// TIA Portal project "PROJECT_PC_SUT" (V17)

(* hardware
DEVICE "S7-1500/ET200MP station_1"  S7-1500 station
   slot 0: "Rail_0"  Rack  6ES7 590-1***0-0AA0
   slot 1: "PLC_2"  CPU 1513-1 PN  6ES7 513-1AL01-0AB0  V2.9
      slot 3: "CPU display_1"  6ES7591-1AA00-0AA0
      slot 32768: "PROFINET interface_1"  X1
         slot 32769: "Port_1"  X1 P1
         slot 32770: "Port_2"  X1 P2
      slot 34817: "Virtual CP interface port_1"  Virtual CP interface port  Virtual CP interface port
DEVICE "HMI_1"  TP700 Comfort
   slot 0: "HMI_1"  TP700 Comfort  6AV2 124-0GC01-0AX0  17.0.0.0
   slot 1: "HMI_RT_1"  TP700 Comfort  6AV2 124-0GC01-0AX0  17.0.0.0
   slot 5: "HMI_1.IE_CP_1"  PROFINET Interface  17.0.0.0
      slot 1: "PROFINET Interface_1"  PROFINET Interface
         slot 1: "Port_1"  Port
         slot 2: "Port_2"  Port
   slot 7: "HMI_1.MPI/DP_CP_1"  MPI/DP Interface  17.0.0.0
DEVICE "PC-System_1"  SIMATIC PC station
   slot 0: "SIMATIC PC station"  Rail  SIMATIC PC-Station  V1.0
      slot 125: "Stationmanager"  Station_Manager  V6.0.4
   slot 1: "IE general_1"  IE General  IE_CP  V8.2.0
      slot 1: "PROFINET interface"  IEGeneral.Interface.8.2.0
   slot 2: "HMI_RT_2"  WinCC RT Advanced  6AV2 104-0xxxx-xxxx  17.0.0.0
      slot 33792: "Computer interface"  Host interface
*)

// ===== PLC "PLC_2"  CPU 1513-1 PN =====

VAR_GLOBAL   // PLC tag table "Tag_Table"
   "start" AT %I0.1 : Bool;
   "AI1_level_sensor" AT %IW1 : Int;
   "AI2_temp_sensor" AT %IW3 : Int;
   "set_temperature_MW4" AT %MW4 : Int;
   "initial_temperature_MW6" AT %MW6 : Int;
   "set_level_MW2" AT %MW2 : Int;
   "gain" AT %MW8 : Int;
   "valve1" AT %Q0.1 : Bool;
   "valve2" AT %Q0.2 : Bool;
   "valve3" AT %Q0.3 : Bool;
   "valve4" AT %Q0.4 : Bool;
   "valve5" AT %Q0.5 : Bool;
   "mixer_motor" AT %Q0.6 : Bool;
   "AV1" AT %QW2 : Word;
   "AV2" AT %QW4 : Int;
   "compare_level" AT %MD10 : Real;
   "flag1" AT %M22.0 : Bool;
   "compare_bit_for_heating" AT %M22.1 : Bool;
   "set_heating" AT %M22.2 : Bool;
   "flag2" AT %M22.3 : Bool;
   "flag3" AT %M22.4 : Bool;
   "set_cooling" AT %M22.5 : Bool;
   "flag0" AT %M22.6 : Bool;
   "compare_bit_reset" AT %M22.7 : Bool;
   "compare_drain_bit_1" AT %M23.0 : Bool;
   "compare_drain_bit_2" AT %M23.1 : Bool;
   "drain_activation_bit" AT %M23.2 : Bool;
END_VAR

// folder: System blocks/Program resources

DATA_BLOCK "Timer_1"   // DB1
{ S7_Optimized_Access := 'TRUE' }
AUTHOR : Simatic
FAMILY : IEC
NAME : IEC_TMR
VERSION : 1.0
// stored: InstanceOfName IEC_TIMER
"IEC_TIMER"
BEGIN
END_DATA_BLOCK

// folder: (top level)

FUNCTION "compare_level_value" : Void   // FC1, LAD
{ S7_Optimized_Access := 'TRUE' }
VERSION : 0.1
   VAR_INPUT
      set_level_MW2 : Int;
   END_VAR
   VAR_OUTPUT
      compare_level : Real;
   END_VAR
   VAR_TEMP
      hold : Real;
      set_level_convert : Real;
   END_VAR
BEGIN

REGION Network 1: Data type conversion
   // covert set_level_MW2 from INT to REAL
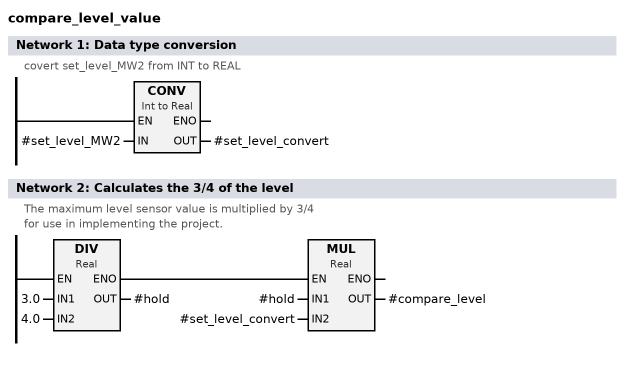
   RUNG wire#powerrail
      { S7_Templates := "[SrcType := Int, DestType := Real]" } Convert(in := #set_level_MW2, out => #set_level_convert)
   END_RUNG
   // the same network as SCL:
   #set_level_convert := INT_TO_REAL(#set_level_MW2);
END_REGION

REGION Network 2: Calculates the 3/4 of the level
   // The maximum level sensor value is multiplied by 3/4
   // for use in implementing the project.
   RUNG wire#powerrail
      { S7_Templates := "SrcType := Real" } Div(in1 := 3.0, in2 := 4.0, out => #hold)
      { S7_Templates := "SrcType := Real" } Mul(in1 := #hold, in2 := #set_level_convert, out => #compare_level)
   END_RUNG
   // the same network as SCL:
   #hold := 3.0 / 4.0;
   #compare_level := #hold * #set_level_convert;
END_REGION
END_FUNCTION

FUNCTION "Filling" : Void   // FC2, LAD
{ S7_Optimized_Access := 'TRUE' }
VERSION : 0.1
   VAR_INPUT
      valve3 : Bool;
      valve4 : Bool;
      valve5 : Bool;
      AI1_level_sensor : Int;
      compare_level : Real;
      set_level_MW2 : Int;
   END_VAR
   VAR_OUTPUT
      valve1 : Bool;
      valve2 : Bool;
      mixer_motor : Bool;
      flag0 : Bool;
   END_VAR
   VAR_TEMP
      level_sensor_conv : Real;
      set_level_converted : Real;
   END_VAR
   VAR_TEMP   // added for the SCL form of the ladder/FBD networks
      _w1 : Bool;
   END_VAR
BEGIN

REGION Network 1: Data type convert
   // A1I_level_sensor data type is converted to Real
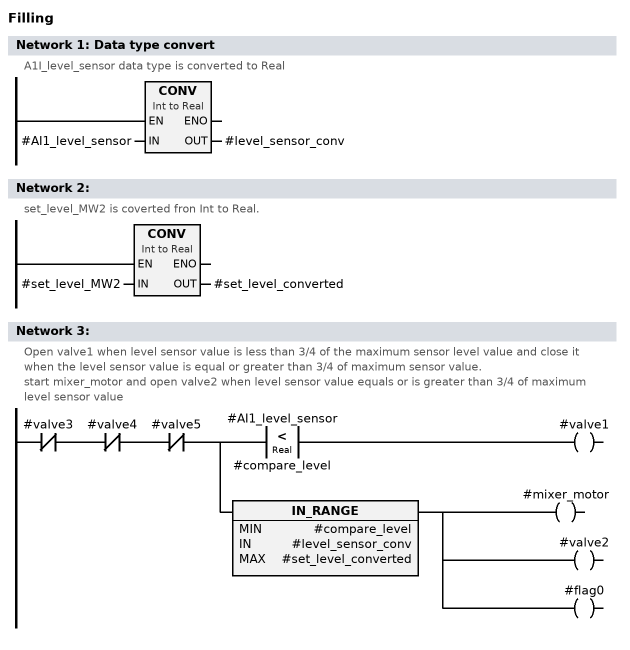
   RUNG wire#powerrail
      { S7_Templates := "[SrcType := Int, DestType := Real]" } Convert(in := #AI1_level_sensor, out => #level_sensor_conv)
   END_RUNG
   // the same network as SCL:
   #level_sensor_conv := INT_TO_REAL(#AI1_level_sensor);
END_REGION

REGION Network 2
   // set_level_MW2 is coverted fron Int to Real.
   RUNG wire#powerrail
      { S7_Templates := "[SrcType := Int, DestType := Real]" } Convert(in := #set_level_MW2, out => #set_level_converted)
   END_RUNG
   // the same network as SCL:
   #set_level_converted := INT_TO_REAL(#set_level_MW2);
END_REGION

REGION Network 3
   // Open valve1 when level sensor value is less than 3/4 of the maximum sensor level value and close it when the level sensor value is equal or greater than 3/4 of maximum sensor value.
   // 
   // start mixer_motor and open valve2 when level sensor value equals or is greater than 3/4 of maximum level sensor value
   RUNG wire#powerrail
      I_Contact( #valve3 )
      I_Contact( #valve4 )
      I_Contact( #valve5 )
      wire#w1
      { S7_Templates := "SrcType := Real" } LT_Contact(in1 := #AI1_level_sensor, in2 := #compare_level)
      Coil( #valve1 )
   END_RUNG
   RUNG wire#w1
      { S7_Templates := "SrcType := Real" } InRange(min := #compare_level, in := #level_sensor_conv, max := #set_level_converted)
      wire#w2
      Coil( #mixer_motor )
   END_RUNG
   RUNG wire#w2
      Coil( #valve2 )
   END_RUNG
   RUNG wire#w2
      Coil( #flag0 )
   END_RUNG
   // the same network as SCL:
   #_w1 := NOT #valve3 AND NOT #valve4 AND NOT #valve5;
   #valve1 := #_w1 AND (#AI1_level_sensor < #compare_level);
   #mixer_motor := #_w1 AND (#compare_level <= #level_sensor_conv) AND (#level_sensor_conv <= #set_level_converted);
   #valve2 := #mixer_motor;
   #flag0 := #mixer_motor;
END_REGION
END_FUNCTION

FUNCTION "P_Controller" : Void   // FC3, LAD
{ S7_Optimized_Access := 'TRUE' }
VERSION : 0.1
// Proportional controller for the system
   VAR_INPUT
      AI2_temp_sensor : Int;
      gain : Int;
      set_temperature_MW4 : Int;
   END_VAR
   VAR_OUTPUT
      AV2 : Int;
   END_VAR
   VAR_TEMP
      error : Int;
      multiply : Real;
      norm_out : Real;
      limit_out : Real;
   END_VAR
BEGIN

REGION Network 1
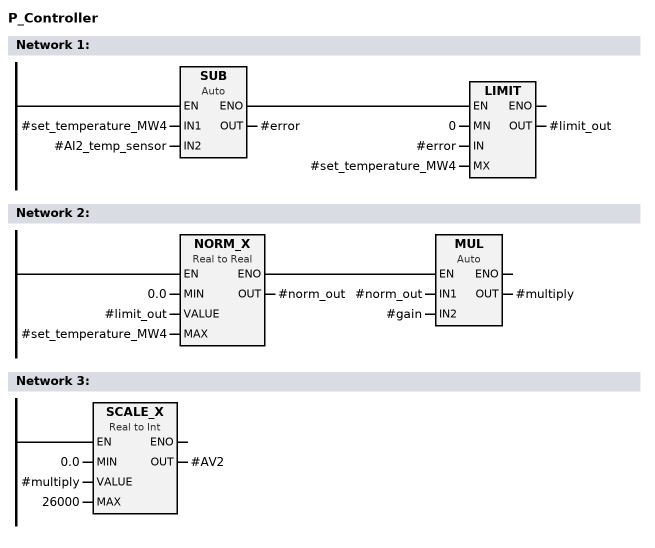
   #error := #set_temperature_MW4 - #AI2_temp_sensor;
   #limit_out := LIMIT(MN := 0, IN := #error, MX := #set_temperature_MW4);
END_REGION

REGION Network 2
   RUNG wire#powerrail
      { S7_Templates := "[SrcType := Real, DestType := Real]" } Normalize(min := 0.0, value := #limit_out, max := #set_temperature_MW4, out => #norm_out)
      Mul(in1 := #norm_out, in2 := #gain, out => #multiply)
   END_RUNG
   // the same network as SCL:
   #norm_out := NORM_X(MIN := 0.0, VALUE := #limit_out, MAX := #set_temperature_MW4);
   #multiply := #norm_out * #gain;
END_REGION

REGION Network 3
   RUNG wire#powerrail
      { S7_Templates := "[SrcType := Real, DestType := Int]" } Scale(min := 0.0, value := #multiply, max := 26000, out => #AV2)
   END_RUNG
   // the same network as SCL:
   #AV2 := SCALE_X(MIN := 0.0, VALUE := #multiply, MAX := 26000);
END_REGION
END_FUNCTION

FUNCTION "heating" : Void   // FC4, LAD
{ S7_Optimized_Access := 'TRUE' }
VERSION : 0.1
   VAR_INPUT
      AI2_temp_sensor : Int;
      valve3 : Bool;
      valve4 : Bool;
      set_temperture_MW4 : Int;
      gain : Int;
   END_VAR
   VAR_OUTPUT
      valve5 : Bool;
      AV2 : Int;
   END_VAR
   VAR_IN_OUT
      trigger_move : Bool;
      flag1 : Bool;
   END_VAR
   VAR_TEMP
      bit_operate : Bool;
   END_VAR
BEGIN

REGION Network 1
   // Reset flag1, which stops mixer_motor and closes valve2 when level sensor value is greater than the set_level sensor value.
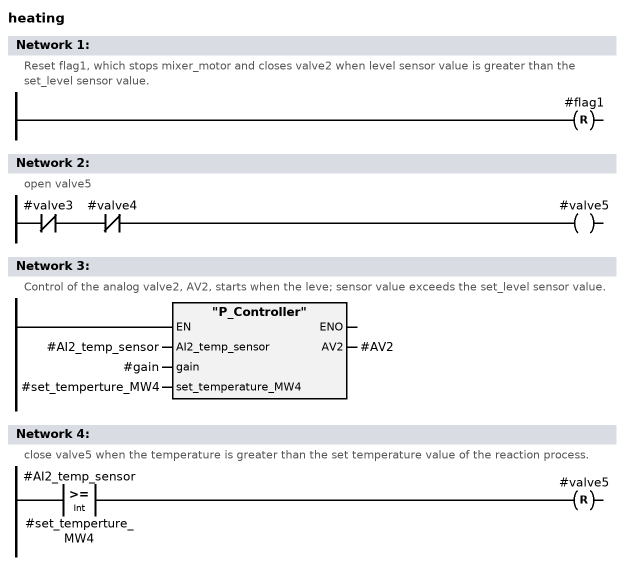
   RUNG wire#powerrail
      R_Coil( #flag1 )
   END_RUNG
   // the same network as SCL:
   #flag1 := FALSE;
END_REGION

REGION Network 2
   // open valve5
   RUNG wire#powerrail
      I_Contact( #valve3 )
      I_Contact( #valve4 )
      Coil( #valve5 )
   END_RUNG
   // the same network as SCL:
   #valve5 := NOT #valve3 AND NOT #valve4;
END_REGION

REGION Network 3
   // Control of the analog valve2, AV2, starts when the leve; sensor value exceeds the set_level sensor value.
   RUNG wire#powerrail
      "P_Controller"(AI2_temp_sensor := #AI2_temp_sensor, gain := #gain, set_temperature_MW4 := #set_temperture_MW4, AV2 => #AV2)
   END_RUNG
   // the same network as SCL:
   "P_Controller"(AI2_temp_sensor := #AI2_temp_sensor,
                  gain := #gain,
                  set_temperature_MW4 := #set_temperture_MW4,
                  AV2 => #AV2);
END_REGION

REGION Network 4
   // close valve5 when the temperature is greater than the set temperature value of the reaction process.
   RUNG wire#powerrail
      { S7_Templates := "SrcType := Int" } GE_Contact(in1 := #AI2_temp_sensor, in2 := #set_temperture_MW4)
      R_Coil( #valve5 )
   END_RUNG
   // the same network as SCL:
   IF #AI2_temp_sensor >= #set_temperture_MW4 THEN #valve5 := FALSE; END_IF;
END_REGION
END_FUNCTION

ORGANIZATION_BLOCK "Main"   // OB1, LAD, ProgramCycle
TITLE = "Main Program Sweep (Cycle)"
{ S7_Optimized_Access := 'TRUE' }
VERSION : 0.1
   VAR_INPUT
      Initial_Call : Bool;   // Initial call of this OB
      Remanence : Bool;   // =True, if remanent data are available
   END_VAR
   VAR_TEMP   // added for the SCL form of the ladder/FBD networks
      _w1 : Bool;
      _w2 : Bool;
      _w3 : Bool;
   END_VAR
BEGIN

REGION Network 1: INITIAL STATE OF THE REACTOR
   // In this block, the compare function is called. This compare function is used to control the mixer and filling processes by comparing the level at which the mixer will be turned on and off, and also when the filling valves will be turned on and off.
   // 
   // Also, we set flag1 in this Network, Flag1 will be used to start the filling phase of the process.
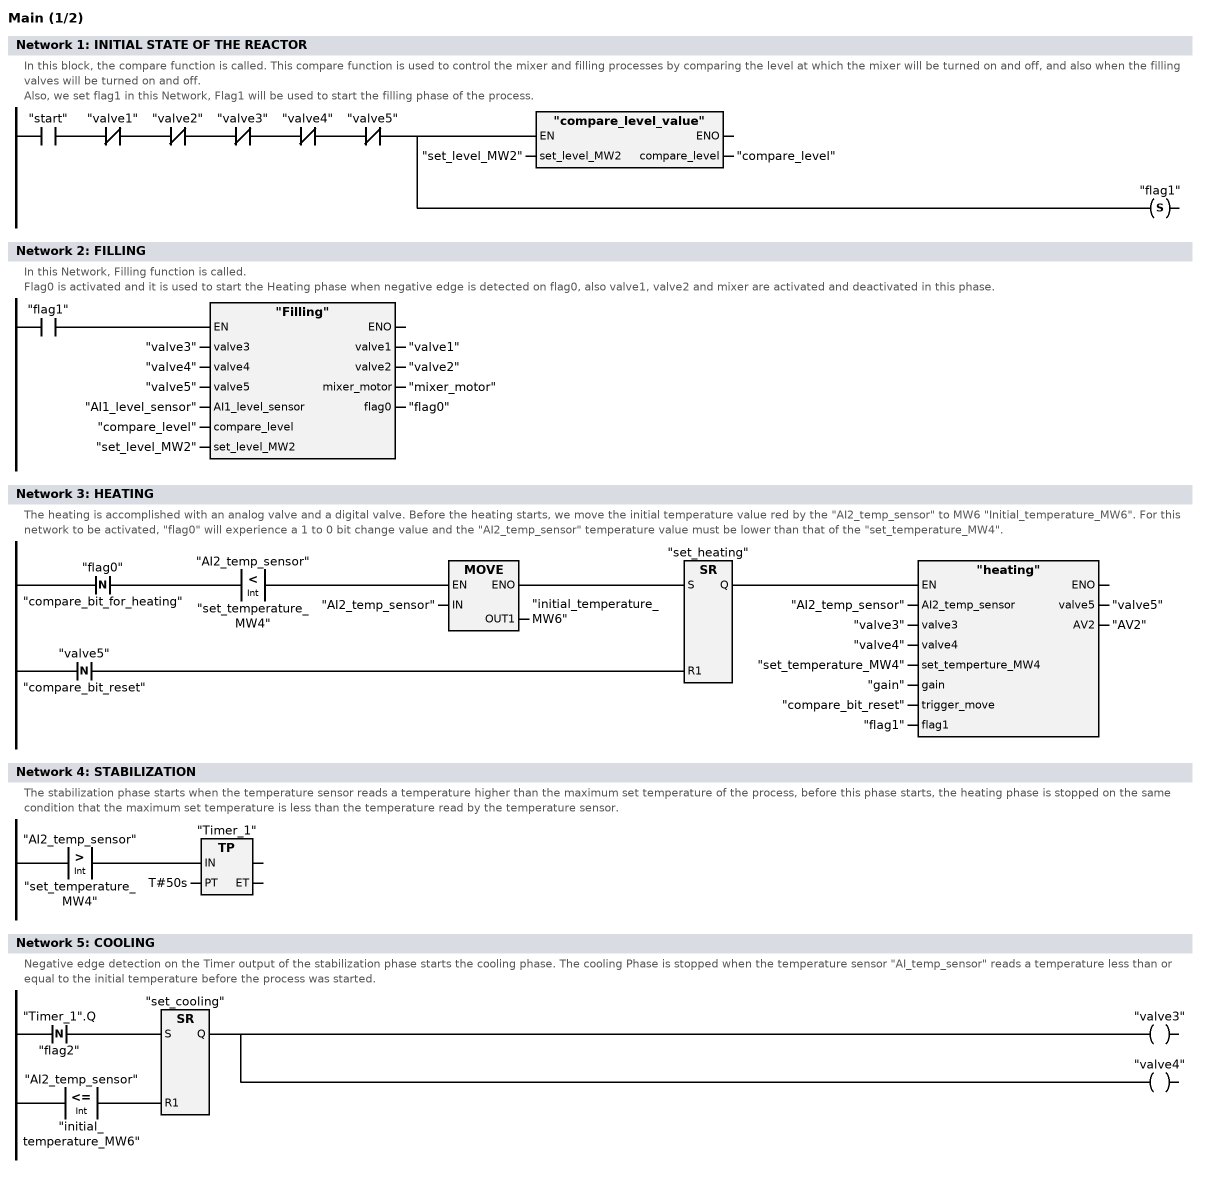
   RUNG wire#powerrail
      Contact( "start" )
      I_Contact( "valve1" )
      I_Contact( "valve2" )
      I_Contact( "valve3" )
      I_Contact( "valve4" )
      I_Contact( "valve5" )
      wire#w1
      "compare_level_value"(set_level_MW2 := "set_level_MW2", compare_level => "compare_level")
   END_RUNG
   RUNG wire#w1
      S_Coil( "flag1" )
   END_RUNG
   // the same network as SCL:
   #_w1 := "start" AND NOT "valve1" AND NOT "valve2" AND NOT "valve3" AND NOT "valve4" AND NOT "valve5";
   IF #_w1 THEN
       "compare_level_value"(set_level_MW2 := "set_level_MW2", compare_level => "compare_level");
       "flag1" := TRUE;
   END_IF;
END_REGION

REGION Network 2: FILLING
   // In this Network, Filling function is called.
   // Flag0 is activated and it is used to start the Heating phase when negative edge is detected on flag0, also valve1, valve2 and mixer are activated and deactivated in this phase.
   RUNG wire#powerrail
      Contact( "flag1" )
      "Filling"(valve3 := "valve3", valve4 := "valve4", valve5 := "valve5", AI1_level_sensor := "AI1_level_sensor", compare_level := "compare_level", set_level_MW2 := "set_level_MW2", valve1 => "valve1", valve2 => "valve2", mixer_motor => "mixer_motor", flag0 => "flag0")
   END_RUNG
   // the same network as SCL:
   IF "flag1" THEN
       "Filling"(valve3 := "valve3",
                 valve4 := "valve4",
                 valve5 := "valve5",
                 AI1_level_sensor := "AI1_level_sensor",
                 compare_level := "compare_level",
                 set_level_MW2 := "set_level_MW2",
                 valve1 => "valve1",
                 valve2 => "valve2",
                 mixer_motor => "mixer_motor",
                 flag0 => "flag0");
   END_IF;
END_REGION

REGION Network 3: HEATING
   // The heating is accomplished with an analog valve and a digital valve. Before the heating starts, we move the initial temperature value red by the "AI2_temp_sensor" to MW6 "Initial_temperature_MW6". For this network to be activated, "flag0" will experience a 1 to 0 bit change value and the "AI2_temp_sensor" temperature value must be lower than that of the "set_temperature_MW4".
   RUNG wire#powerrail
      N_Contact(operand := "flag0", bit := "compare_bit_for_heating")
      { S7_Templates := "SrcType := Int" } LT_Contact(in1 := "AI2_temp_sensor", in2 := "set_temperature_MW4")
      Move(in := "AI2_temp_sensor", out1 => "initial_temperature_MW6")
      S_SR(operand := "set_heating", r1 := wire#w1)
      "heating"(AI2_temp_sensor := "AI2_temp_sensor", valve3 := "valve3", valve4 := "valve4", set_temperture_MW4 := "set_temperature_MW4", gain := "gain", trigger_move := "compare_bit_reset", flag1 := "flag1", valve5 => "valve5", AV2 => "AV2")
   END_RUNG
   RUNG wire#powerrail
      N_Contact(operand := "valve5", bit := "compare_bit_reset")
   END_RUNG wire#w1
   // the same network as SCL:
   #_w1 := NOT "flag0" AND "compare_bit_for_heating";   // falling edge of "flag0"
   "compare_bit_for_heating" := "flag0";
   #_w2 := #_w1 AND ("AI2_temp_sensor" < "set_temperature_MW4");
   IF #_w2 THEN "initial_temperature_MW6" := "AI2_temp_sensor"; END_IF;
   #_w3 := NOT "valve5" AND "compare_bit_reset";   // falling edge of "valve5"
   "compare_bit_reset" := "valve5";
   IF #_w2 THEN
       "set_heating" := TRUE;   // SR flip-flop
   END_IF;
   IF #_w3 THEN "set_heating" := FALSE; END_IF;
   IF "set_heating" THEN
       "heating"(AI2_temp_sensor := "AI2_temp_sensor",
                 valve3 := "valve3",
                 valve4 := "valve4",
                 set_temperture_MW4 := "set_temperature_MW4",
                 gain := "gain",
                 trigger_move := "compare_bit_reset",
                 flag1 := "flag1",
                 valve5 => "valve5",
                 AV2 => "AV2");
   END_IF;
END_REGION

REGION Network 4: STABILIZATION
   // The stabilization phase starts when the temperature sensor reads a temperature higher than the maximum set temperature of the process, before this phase starts, the heating phase is stopped on the same condition that the maximum set temperature is less than the temperature read by the temperature sensor.
   "Timer_1".TP(IN := "AI2_temp_sensor" > "set_temperature_MW4", PT := T#50s);
END_REGION

REGION Network 5: COOLING
   // Negative edge detection on the Timer output of the stabilization phase starts the cooling phase. The cooling Phase is stopped when the temperature sensor "AI_temp_sensor" reads a temperature less than or equal to the initial temperature before the process was started.
   RUNG wire#powerrail
      N_Contact(operand := "Timer_1".Q, bit := "flag2")
      S_SR(operand := "set_cooling", r1 := wire#w1)
      wire#w2
      Coil( "valve3" )
   END_RUNG
   RUNG wire#powerrail
      { S7_Templates := "SrcType := Int" } LE_Contact(in1 := "AI2_temp_sensor", in2 := "initial_temperature_MW6")
   END_RUNG wire#w1
   RUNG wire#w2
      Coil( "valve4" )
   END_RUNG
   // the same network as SCL:
   #_w1 := NOT "Timer_1".Q AND "flag2";   // falling edge of "Timer_1".Q
   "flag2" := "Timer_1".Q;
   IF #_w1 THEN
       "set_cooling" := TRUE;   // SR flip-flop
   END_IF;
   IF "AI2_temp_sensor" <= "initial_temperature_MW6" THEN "set_cooling" := FALSE; END_IF;
   "valve3" := "set_cooling";
   "valve4" := "set_cooling";
END_REGION

REGION Network 6: DRAINING
   // This phase is started when the cooling valves experiences a 1 to 0 bit change and the level sensor reads a level above 20litres.
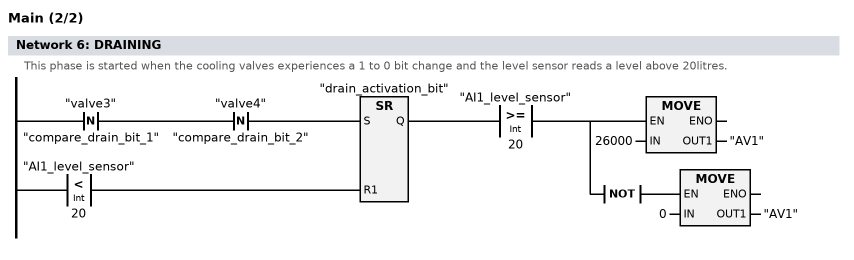
   RUNG wire#powerrail
      N_Contact(operand := "valve3", bit := "compare_drain_bit_1")
      N_Contact(operand := "valve4", bit := "compare_drain_bit_2")
      S_SR(operand := "drain_activation_bit", r1 := wire#w1)
      { S7_Templates := "SrcType := Int" } GE_Contact(in1 := "AI1_level_sensor", in2 := 20)
      wire#w2
      Move(in := 26000, out1 => "AV1")
   END_RUNG
   RUNG wire#powerrail
      { S7_Templates := "SrcType := Int" } LT_Contact(in1 := "AI1_level_sensor", in2 := 20)
   END_RUNG wire#w1
   RUNG wire#w2
      Not()
      Move(in := 0, out1 => "AV1")
   END_RUNG
   // the same network as SCL:
   #_w1 := NOT "valve3" AND "compare_drain_bit_1";   // falling edge of "valve3"
   "compare_drain_bit_1" := "valve3";
   #_w2 := #_w1 AND NOT "valve4" AND "compare_drain_bit_2";   // falling edge of "valve4"
   "compare_drain_bit_2" := "valve4";
   IF #_w2 THEN
       "drain_activation_bit" := TRUE;   // SR flip-flop
   END_IF;
   IF "AI1_level_sensor" < 20 THEN "drain_activation_bit" := FALSE; END_IF;
   #_w3 := "drain_activation_bit" AND ("AI1_level_sensor" >= 20);
   IF #_w3 THEN "AV1" := 26000; END_IF;
   IF NOT #_w3 THEN "AV1" := 0; END_IF;
END_REGION
END_ORGANIZATION_BLOCK

(* ===== HMI "HMI_RT_1" =====
connection "HMI_Connection_1": ETHERNET, S7_1500_OMS

HMI tags "Default tag table"
   "HMI_AI_level" : Int = PLC AI1_level_sensor AT %IW1, 1 s
   "HMI_gain" : Int = PLC gain AT %MW8, 1 s
   "HMI_set" : Int = PLC set_temperature_MW4 AT %MW4, 1 s
   "HMI_AV2" : Int = PLC AV2 AT %QW4, 1 s
   "HMI_A2_temperature_sensor" : Int = PLC AI2_temp_sensor AT %IW3, 1 s

screen "Screen_1" 800x480
   IOField "I/O field_1" at 8,33 size 158x48; FormatPattern s99999
      ProcessValue <- "HMI_AI_level"
   IOField "I/O field_2" at 585,30 size 149x48; FormatPattern s99999
      ProcessValue <- "HMI_AV2"
   IOField "I/O field_3" at 8,232 size 147x37; FormatPattern s99999
      ProcessValue <- "HMI_A2_temperature_sensor"
   IOField "I/O field_4" at 8,302 size 147x42; FormatPattern s99999
      ProcessValue <- "HMI_set"
   IOField "I/O field_5" at 8,155 size 147x37; FormatPattern s99999
      ProcessValue <- "HMI_gain"
   TextField "Text field_1" at 17,7 size 114x23; Text 'level sensor'
   TextField "Text field_2" at 10,129 size 46x23; Text 'Gain'
   TextField "Text field_3" at 9,209 size 120x23; Text 'Temp sensor'
   TextField "Text field_4" at 9,281 size 91x23; Text 'Set Temp'
   TextField "Text field_5" at 581,5 size 124x23; Text 'Analog Valve'
*)